FUNCTION_BLOCK "FB_CrossCutsModbus_V1.00"   // FB1, LAD
TITLE = Cross cut machine V1.00
{ S7_Optimized_Access := 'TRUE' }
VERSION : 0.1
   VAR_INPUT
      IN_dMachineIndex : DInt;   // Tracking machine index
      IN_dGlassBreakMachineIndex : DInt;   // Glass break machine index
      IN_dGlassSearchMachineIndex_Q0 : DInt;   // Glass search machine index
      IN_dGlassSearchMachineIndex_Q1 : DInt;   // Glass search machine index
      IN_dGlassSearchMachineIndex_Q2 : DInt;   // Glass search machine index
      IN_dGlassSearchMachineIndex_Q3 : DInt;   // Glass search machine index
      IN_dXCutIndex : DInt;   // Index of the XCUT (0=XC#1, 1=XC#2...)
      IN_xCycleON : Bool;   // Cycle ON
      IN_xGeneralReset : Bool;   // General reset
      IN_xResetAlarms : Bool;   // Reset alarms
      IN_xFaultsEnabled : Bool;   // Faults enabled
      IN_xSimulationActive : Bool;   // Enable simulation (EXPERT USER)
      IN_xMBDone : Bool;   // Modbus client done
      IN_xMBError : Bool;   // Xcut DB
   END_VAR
   VAR_IN_OUT
      INO_tTrack : "UDT_CapData_Tracking";   // Tracking plate
      INO_tEnc : "UDT_Encoder";   // Encoder data
      INO_tOBInit : "GP_OB_Initialize";   // OB Initialize
      INO_tRibbon : "UDT_RibbonData";   // Ribbon data
      INO_tXCutOpt : "FB_CrossCutOpt_V1.00";   // Ribbon data
   END_VAR
   VAR RETAIN
      tHMW : Struct   // HMI Write data
         xCutBreakEnabled : Bool;   // Cut on glass break enabled {X|X|X|X|O}
         xUpdateDistSnap : Bool;   // Update distance from snap roll {X|X|X|X|M}
         xUpdateAngleValue : Bool;   // Update angle value {X|X|X|X|M}
         xIncAngleValue : Bool;   // Increment angle value {X|X|X|X|O}
         xDecAngleValue : Bool;   // Decrement angle value {X|X|X|X|O}
         xUpdateDistCenterLine : Bool;   // Update distance from center line {X|X|X|X|M}
         xCalibDistRequest : Bool;   // Calibration distance request {X|X|X|X|O}
         xCalibDiagRequest : Bool;   // Calibration diagonal request {X|X|X|X|O}
         tManCmd : Struct   // Manual command
            xMan_JogForward : Bool;   // Manual mode - Jog forward {X|X|X|X|M}
            xMan_JobBackward : Bool;   // Manual mode - Jog backward {X|X|X|X|M}
            xMan_CarriageDown : Bool;   // Manual mode - Carriage down {X|X|X|X|M}
            xMan_FireOn : Bool;   // Manual mode - Fire ON {X|X|X|X|M}
            xMan_OilOn : Bool;   // Manual mode - Oil ON {X|X|X|X|M}
         END_STRUCT;
         xCutOperator : Bool;   // Cutting position by operator request {X|X|X|X|O}
         xCutGross : Bool;   // Cutting position by gross width position {X|X|X|X|O}
         xCutNet : Bool;   // Cutting position by net width position {X|X|X|X|O}
         xCutYCut : Bool;   // Cutting position by YCut position {X|X|X|X|O}
         dOperStartCutPos_cmm : DInt;   // Operator start cut position [mm/100] {mm/100|mm|-3000|0|O}
         dOperEndCutPos_cmm : DInt;   // Operator end cut position [mm/100] {mm/100|mm|0|3000|O}
         dDescReactTime_ms : DInt;   // Carriage descent reaction time [ms] {ms|s|0|1|M}
         dRaiseReactTime_ms : DInt;   // Carriage raise reaction time [ms] {ms|s|0|1|M}
         dFireONReactTime_ms : DInt;   // Fire ON reaction time [ms] {ms|s|0|1|M}
         dFireOFFReactTime_ms : DInt;   // Fire OFF reaction time [ms] {ms|s|0|1|M}
         dOilONDelay_ms : DInt;   // Oil ON delay [ms] {ms|s|-1|1|O}
         dOilOFFDelay_ms : DInt;   // Oil OFF delay [ms] {ms|s|-1|1|O}
         dCutStartOffsetDelay_cmm : DInt;   // Start cut offset delay [mm/100] {mm/100|mm|-500|500|O}
         dCutEndOffsetDelay_cmm : DInt;   // End cut offset delay [mm/100] {mm/100|mm|-500|500|O}
         dDistanceFromSnaproll_cmm : DInt;   // Distance from snaproll [mm/100] {mm/100|mm|0|10000|M}
         dAngleValue_uDegree : DInt;   // Bridge angle value [°/1000000] {°/1000000|°|7|9|M}
         dDistanceFromCenterLine_cmm : DInt;   // Distance from center line [mm/100] {mm/100|mm|-3000|0|M}
         dDistTeoLength_cmm : DInt;   // Calibration distance.Theorical length [mm/100] {mm/100|mm|0|7000|O}
         dDistRealLength_cmm : DInt;   // Calibration distance.Real length [mm/100] {mm/100|mm|0|7000|O}
         dDiagRealLength_cmm : DInt;   // Calibration diagonal.Real length [mm/100] {mm/100|mm|0|7000|O}
         dDiagRealWidth_cmm : DInt;   // Calibration diagonal.Real width [mm/100] {mm/100|mm|0|4000|O}
         dDiagGlassFlow_cmm : DInt;   // Calibration diagonal.Real length diagonal glass flow [mm/100] {mm/100|mm|0|10000|O}
         dDiagGlassOppFlow_cmm : DInt;   // Calibration diagonal.Real length diagonal opposite glass flow [mm/100] {mm/100|mm|0|10000|O}
         dCuttingPressure_mN : DInt;   // Cutting pressure [N/1000] {N/1000|N|9|180|O}
         dPosOffset_cmm : DInt;   // Calibration offset distance from snaproll [mm/100] {mm/100|mm|-50|50|O}
         dCutPriority : DInt;   // Cut priority number {X|X|0|5|O}
         xResetHeadUsage : Bool;   // Reset the head usage {X|X|X|X|O}
         xEnDisManCom : Bool;   // Enable disable manual command {X|X|X|X|M}
      END_STRUCT;
      tHMR : Struct   // HMI Read data
         tManCmd : Struct   // Manual command
            xManJogFwdFdbk : Bool;   // Manual jog forward feedback {X|X|X|X|O}
            xManJogBckFdbk : Bool;   // Manual jog backward feedback {X|X|X|X|O}
            xManCarriageDownFdbk : Bool;   // Manual carriage down feedback {X|X|X|X|O}
            xManFireONFdbk : Bool;   // Manual fire ON feedback {X|X|X|X|O}
            xManOilONFdbk : Bool;   // Manual oil ON feedback {X|X|X|X|O}
         END_STRUCT;
         dActualCutPosRequest : DInt;   // Actual cut position request (1=By operator 2=On gross ribbon 3=On net ribbon 4=On YCut position) {X|X|X|X|O}
         dXCutStatusRequest : DInt;   // XCut status request (1=Disabled 3=Enabled) {X|X|X|X|O}
         dXCutActualStatus : DInt;   // XCut actual status (1=Disabled 3=Enabled) {X|X|X|X|O}
         dDistanceFromSnaproll_cmm : DInt;   // Distance from snaproll [mm/100] {mm/100|mm|X|X|O}
         dAngleValue_uDegree : DInt;   // Angle value [°/1000000] {°/1000000|°|X|X|O}
         dDistanceFromCenterLine_cmm : DInt;   // Distance from center line [mm/100] {mm/100|mm|X|X|O}
         dCarriagePosition_cmm : DInt;   // Actual carriage position [mm/100]
         dStatus : DInt;   // XCut actual status (1=Idle 3=Running 7=Faulted) {X|X|X|X|O}
         rHeadUsage_km : Real;   // Head usage [Km] {Km|Km|X|X|O}
         xManComEn : Bool;   // Manual command enabled {X|X|X|X|O}
         dTimeHeadDown_ms : DInt;   // Time head down [ms] {ms|s|X|X|O}
      END_STRUCT;
   END_VAR
   VAR
      tALM : Struct   // HMI Alarms
         tE : Struct   // Emergency alarms
            xLocON : Bool;   // KE.Local emergency ON {X|X|X|X|O}
            xLocal1 : Bool;   // SB.Local emergency push button 1 {X|X|X|X|O}
            xLocal2 : Bool;   // SB.Local emergency push button 2 {X|X|X|X|O}
            xLocal3 : Bool;   // SB.Local emergency push button 3 {X|X|X|X|O}
            xSpare_4 : Bool;
            xSpare_5 : Bool;
            xSpare_6 : Bool;
            xSpare_7 : Bool;
            xSpare_8 : Bool;
            xSpare_9 : Bool;
            xSpare_10 : Bool;
            xSpare_11 : Bool;
            xSpare_12 : Bool;
            xSpare_13 : Bool;
            xSpare_14 : Bool;
            xSpare_15 : Bool;
            xSpare_16 : Bool;
            xSpare_17 : Bool;
            xSpare_18 : Bool;
            xSpare_19 : Bool;
            xSpare_20 : Bool;
            xSpare_21 : Bool;
            xSpare_22 : Bool;
            xSpare_23 : Bool;
            xSpare_24 : Bool;
            xSpare_25 : Bool;
            xSpare_26 : Bool;
            xSpare_27 : Bool;
            xSpare_28 : Bool;
            xSpare_29 : Bool;
            xSpare_30 : Bool;
            xSpare_31 : Bool;
         END_STRUCT;
         tS : Struct   // Stopping faults
            xAxisNotAvail : Bool;   // AZ.Axis not available {X|X|X|X|O}
            xInpInstallation : Bool;   // L+.Input power supply ON {X|X|X|X|O}
            xAuxPower : Bool;   // L+.Auxiliary power supple set-in {X|X|X|X|O}
            xAreaSafety : Bool;   // KE.Area safety {X|X|X|X|O}
            xOverstroke : Bool;   // KA.Carriage overstroke {X|X|X|X|O}
            xExternInputPower : Bool;   // L+.External input power supply {X|X|X|X|O}
            xCarriageCutOut : Bool;   // QM.Carriage translation overload {X|X|X|X|O}
            xDriveTrip : Bool;   // AZ.Drive trip {X|X|X|X|O}
            xDriveNotEnabled : Bool;   // AZ.Drive not enabled {X|X|X|X|O}
            xAxisNotReady : Bool;   // AZ.Axis not ready {X|X|X|X|O}
            xDriveNotReady : Bool;   // AZ.Drive not ready {X|X|X|X|O}
            xAxisNotSyncro : Bool;   // AZ.Axis not syncronized {X|X|X|X|O}
            xSpare_12 : Bool;
            xSpare_13 : Bool;
            xSpare_14 : Bool;
            xSpare_15 : Bool;
            xSpare_16 : Bool;
            xSpare_17 : Bool;
            xSpare_18 : Bool;
            xSpare_19 : Bool;
            xSpare_20 : Bool;
            xSpare_21 : Bool;
            xSpare_22 : Bool;
            xSpare_23 : Bool;
            xSpare_24 : Bool;
            xSpare_25 : Bool;
            xSpare_26 : Bool;
            xSpare_27 : Bool;
            xSpare_28 : Bool;
            xSpare_29 : Bool;
            xSpare_30 : Bool;
            xSpare_31 : Bool;
         END_STRUCT;
         tF : Struct   // Faults
            xSpare_0 : Bool;
            xSpare_1 : Bool;
            xSpare_2 : Bool;
            xSpare_3 : Bool;
            xSpare_4 : Bool;
            xSpare_5 : Bool;
            xSpare_6 : Bool;
            xSpare_7 : Bool;
            xSpare_8 : Bool;
            xSpare_9 : Bool;
            xSpare_10 : Bool;
            xSpare_11 : Bool;
            xSpare_12 : Bool;
            xSpare_13 : Bool;
            xSpare_14 : Bool;
            xSpare_15 : Bool;
            xSpare_16 : Bool;
            xSpare_17 : Bool;
            xSpare_18 : Bool;
            xSpare_19 : Bool;
            xSpare_20 : Bool;
            xSpare_21 : Bool;
            xSpare_22 : Bool;
            xSpare_23 : Bool;
            xSpare_24 : Bool;
            xSpare_25 : Bool;
            xSpare_26 : Bool;
            xSpare_27 : Bool;
            xSpare_28 : Bool;
            xSpare_29 : Bool;
            xSpare_30 : Bool;
            xSpare_31 : Bool;
         END_STRUCT;
         tW : Struct   // Warnings
            xSpare_0 : Bool;
            xSpare_1 : Bool;
            xSpare_2 : Bool;
            xSpare_3 : Bool;
            xSpare_4 : Bool;
            xSpare_5 : Bool;
            xSpare_6 : Bool;
            xSpare_7 : Bool;
            xSpare_8 : Bool;
            xSpare_9 : Bool;
            xSpare_10 : Bool;
            xSpare_11 : Bool;
            xSpare_12 : Bool;
            xSpare_13 : Bool;
            xSpare_14 : Bool;
            xSpare_15 : Bool;
            xSpare_16 : Bool;
            xSpare_17 : Bool;
            xSpare_18 : Bool;
            xSpare_19 : Bool;
            xSpare_20 : Bool;
            xSpare_21 : Bool;
            xSpare_22 : Bool;
            xSpare_23 : Bool;
            xSpare_24 : Bool;
            xSpare_25 : Bool;
            xSpare_26 : Bool;
            xSpare_27 : Bool;
            xSpare_28 : Bool;
            xSpare_29 : Bool;
            xSpare_30 : Bool;
            xSpare_31 : Bool;
         END_STRUCT;
      END_STRUCT;
      ST_xPhaseInProgress : Bool;   // Phases are in progress
      AUX_xValidUpCap : Bool;   // Upstream cap is valid
      AUX_xValidDwCap : Bool;   // Downstream cap is valid
      AUX_dUpCapIndex : DInt;   // Index of the upstream cap
      AUX_dDwCapIndex : DInt;   // Index of the downstream cap
      OS_xNewCapUp : Bool;   // New cap arrived upstream
      OS_xNewCapDw : Bool;   // New cap arrived downstream
      OS_xNewCap : Bool;   // New cap arrived
      ST_xStoppingFaults : Bool;   // Stopping faults
      ST_xFaults : Bool;   // Faults
      ST_xWarnings : Bool;   // Warnings
      ST_xOutputEnabled : Bool;   // Output enabled
      ST_xGlassBreak : Bool;   // Glass break under bridge
      ST_xQualitWithFixedXcut : Bool;   // Quality cap with fixed xcut choice coming
      AUX_dCutStartPosUp_cmm : DInt;   // Cut start position upstream [mm/100]
      AUX_dCutStopPosUp_cmm : DInt;   // Cut stop position downstream [mm/100]
      AUX_dCutStartPosDw_cmm : DInt;   // Cut start position downstream [mm/100]
      AUX_dCutStopPosDw_cmm : DInt;   // Cut stop position downstream [mm/100]
      AUX_xUpIsQuality : Bool;   // Upstream cap is a quality cap
      AUX_xDwIsQuality : Bool;   // Downstream cap is a quality cap
      PH_xCutRequest : Bool;   // Cut request phase
      PH_xWriteModbus : Bool;   // Modbus write phase
      PH_xEndWriteModbus : Bool;   // Modbus end write phase
      PH_xReadModbus : Bool;   // Modbus read phase
      PH_xEndReadModbus : Bool;   // Modbus end read phase
      AUX_dMissionCounterValue_cmm : DInt;   // Mission counter value to inverter [mm/100]
      AUX_dMissionToSend : DInt;   // Index mission send to inverter
      AUX_tOutputDrive : "UDT_XCUT_DRIVE_OUTPUT";   // Copy of output area drive
      PH_xEndCutRequest : Bool;   // End cut request phase
      OSR_xButtonEnabled : Bool;   // OSR.Button enabled
      OS_xButtonEnabled : Bool;   // OS.Button enabled
      AUX_dLastLiveCounter : DInt;
      tmON_InvCoutTimeout : TON_TIME;   // Inverter counter timeout
      tmON_AxisSyncroTimeout : TON_TIME;   // Inverter counter timeout
      AUX_dNextPlateTime_ms : DInt;   // Next plate arriving time [ms]
      AUX_dCutTime20Per_ms : DInt;   // Cutting time at 20 percent [ms]
      AUX_dCutTime40Per_ms : DInt;   // Cutting time at 40 percent [ms]
      AUX_dCutTime60Per_ms : DInt;   // Cutting time at 60 percent [ms]
      AUX_dCutTime80Per_ms : DInt;   // Cutting time at 80 percent [ms]
      AUX_dCutTime100Per_ms : DInt;   // Cutting time at 100 percent [ms]
      ST_xCondOkMan : Bool;   // Condition ok manual command
      AUX_dSimWaitEnd_ms : DInt;   // Simulation waiting end cut [ms]
      AUX_dSimCutTime_ms : DInt;   // Simulation cutting time [ms]
      AUX_dSimCutSpace_cmm : DInt;   // Simulation cutting space [mm/100]
      AUX_dSimStoreCutTime_ms : DInt;   // Simulation saved cutting time [ms]
      AUX_rgdParameterArray : Array[0..39] of DInt;   // Array of xcut parameters (menu 20)
      AUX_rgtIN_tDriveData : "UDT_XCUT_DRIVE_INPUT";   // Drive input data
      AUX_rgtOUT_tDriveData : "UDT_XCUT_DRIVE_OUTPUT";   // Drive output data
   END_VAR
   VAR_TEMP
      TMP_rValue : LReal;   // Temp real value
      TMP_xCalcMission : Bool;   // Temp calculate mission
      TMP_dwValue : DWord;   // Temp Dint value
      TMP_dValue : DInt;   // Temp Dint value
      TMP_xUpdateKM : Bool;   // OS update KM counter
      TMP_dCutTime_ms : DInt;   // Cut time [ms]
      TMP_dConstTime_ms : DInt;   // Const time [ms]
      TMP_rAccTime_s : Real;   // Acceleration time [ms]
      TMP_dTravSpace_cmm : DInt;   // Travel space [mm/100]
      TMP_dCutSpace_cmm : DInt;   // Cut Space [mm/100]
      TMP_dCutYSpace_cmm : DInt;   // Cut y space [mm/100]
      TMP_dConstSpace_cmm : DInt;   // Const space [mm/100]
      TMP_dRampSpace_cmm : DInt;   // Ramp space [mm/100]
      TMP_dRetVal : DInt;   // Ramp space [mm/100]
      TMP_rDiagGlassFlow_cmm : Real;
      TMP_rDiagRealWidth_cmm : Real;
      TMP_rDiagRealLength_cmm : Real;
      TMP_iModbus_mode : UDInt;   // Modbus mode (0=read, 1=write)
      TMP_dModbus_address : UDInt;   // Modbus address
      TMP_dModbus_length : UDInt;   // Modbus data length
      TMP_vDataPointer : Variant;
      TMP_dIndex : DInt;
   END_VAR
   VAR CONSTANT
      CONST_DREACTTIMETRACK_MS : DInt := 50;   // Tracking machine reaction time [ms]
      CONST_DMODECUT_OPERATOR : DInt := 1;   // Cut modality - By operator
      CONST_DMODECUT_GROSS : DInt := 2;   // Cut modality - Gross width
      CONST_DMODECUT_NET : DInt := 3;   // Cut modality - Net width
      CONST_DMODECUT_YCUT : DInt := 4;   // Cut modality - YCut
      CONST_DMINCUTRANGE_CMM : DInt := 25000;   // Minimum cutting start position [mm/100]
      CONST_DMAXCUTRANGE_CMM : DInt := 500000;   // Maximum cutting start position [mm/100]
      CONST_DMAXMISSIONNUM : DInt := 1000;   // Maximum number of mission to XCUT
      CONST_DMAXWAITFEEDBACK_CMM : DInt := 20000;   // Waiting space feedback [mm/100]
      CONST_DDISABLED : DInt := 1;   // Disabled
      CONST_DENABLED : DInt := 3;   // Enabled
      CONST_DSIZEALARMS : UDInt := 32;   // Number of bool on alarms structure
      CONST_DTIMEOUTINVERTER_MS : Time := T#2000ms;   // Inverter counter timeout
      CONST_DMAXRETSPEED_RPM : DInt := 3750;   // Maximum return speed [rpm]
      CONST_DSPEED_CMM_S : DInt := 500000;   // Return travel speed [mm/100/s]
      CONST_DRAMP_CMM_S2 : DInt := 1200000;   // Return travel ramp [mm/100/s]
      CONST_DBREAKDOWNOFF_CMM : DInt := 50000;   // Break downstream offset [mm/100]
      CONST_DBREAKUPOFF_CMM : DInt := 50000;   // Break upstream offset [mm/100]
      CONST_DADDRESSMENU_READ : UDInt := 2001;   // Parameter menu start (#20.01=2001)
      CONST_DADDRESSMENU_WRITE : UDInt := 2010;   // Parameter menu start (#20.01=2001)
      CONST_DSEARCHQLTUPSTREAM_CMM : DInt := 1000000;   // Search qlt cap upstream limit [mm/100]
      CONST_DSEARCHQLTDOWNSTREAM_CMM : DInt := 400000;   // Search qlt cap downstream limit [mm/100]
   END_VAR
   VAR_TEMP   // added for the SCL form of the ladder/FBD networks
      _w1 : Bool;
   END_VAR
   // // AUX_rgdParameterArray[0] : #20.01
   // // AUX_rgdParameterArray[1] : #20.02
   // // AUX_rgdParameterArray[2] : #20.03
   // // AUX_rgdParameterArray[3] : #20.04
   // // AUX_rgdParameterArray[4] : #20.05
   // // AUX_rgdParameterArray[5] : #20.06
   // // AUX_rgdParameterArray[6] : #20.07
   // // AUX_rgdParameterArray[7] : #20.08
   // // AUX_rgdParameterArray[8] : #20.09
   // // AUX_rgdParameterArray[9] : #20.10
   // // AUX_rgdParameterArray[10] : #20.11
   // // AUX_rgdParameterArray[11] : #20.12
   // // AUX_rgdParameterArray[12] : #20.13
   // // AUX_rgdParameterArray[13] : #20.14
   // // AUX_rgdParameterArray[14] : #20.15
   // // AUX_rgdParameterArray[15] : #20.16
   // // AUX_rgdParameterArray[16] : #20.17
   // // AUX_rgdParameterArray[17] : #20.18
   // // AUX_rgdParameterArray[18] : #20.19
   // // AUX_rgdParameterArray[19] : #20.20
   // // AUX_rgdParameterArray[20] : #20.21
   // // AUX_rgdParameterArray[21] : #20.22
   // // AUX_rgdParameterArray[22] : #20.23
   // // AUX_rgdParameterArray[23] : #20.24
   // // AUX_rgdParameterArray[24] : #20.25
   // // AUX_rgdParameterArray[25] : #20.26
   // // AUX_rgdParameterArray[26] : #20.27
   // // AUX_rgdParameterArray[27] : #20.28
   // // AUX_rgdParameterArray[28] : #20.29
   // // AUX_rgdParameterArray[29] : #20.30
   // // AUX_rgdParameterArray[30] : #20.31
   // // AUX_rgdParameterArray[31] : #20.32
   // // AUX_rgdParameterArray[32] : #20.33
   // // AUX_rgdParameterArray[33] : #20.34
   // // AUX_rgdParameterArray[34] : #20.35
   // // AUX_rgdParameterArray[35] : #20.36
   // // AUX_rgdParameterArray[36] : #20.37
   // // AUX_rgdParameterArray[37] : #20.38
   // // AUX_rgdParameterArray[38] : #20.39
   // // AUX_rgdParameterArray[39] : #20.40
BEGIN

REGION Network 1: ####_CONSTANTS_####
END_REGION

REGION Network 2: ####_MATCH_####
END_REGION

REGION Network 3 (SCL): Update data from inverter
   IF #PH_xEndReadModbus THEN

   #AUX_rgtIN_tDriveData.dCarriagePos_dmm := #AUX_rgdParameterArray[30];
   #AUX_rgtIN_tDriveData.dLehrPosition_cmm := #AUX_rgdParameterArray[32];
   #AUX_rgtIN_tDriveData.dLehrSpeed_cmm_min := #AUX_rgdParameterArray[36];
   #AUX_rgtIN_tDriveData.dErrorCode := #AUX_rgdParameterArray[34];
   #AUX_rgtIN_tDriveData.dMissionDone := #AUX_rgdParameterArray[35];
   #AUX_rgtIN_tDriveData.dMissionUnDone := #AUX_rgdParameterArray[33];
   #AUX_rgtIN_tDriveData.iLiveCounter := DINT_TO_INT(#AUX_rgdParameterArray[9]);
   #AUX_rgtIN_tDriveData.iTimeHeadDown_ms := DINT_TO_INT(#AUX_rgdParameterArray[10]);
   #TMP_dwValue := DINT_TO_DWORD(#AUX_rgdParameterArray[29]);
   SCATTER(IN:=#TMP_dwValue,
           OUT=>#AUX_rgtIN_tDriveData.rgxStatusBits);

   #PH_xEndReadModbus := 0;
   END_IF;
END_REGION

REGION Network 4 (SCL): General reset
   IF #IN_xGeneralReset THEN

       #PH_xCutRequest := FALSE;
       #PH_xEndCutRequest := FALSE;
       #AUX_xValidDwCap := FALSE;
       #AUX_xValidUpCap := FALSE;

   END_IF;
END_REGION

REGION Network 5 (SCL): Move data information to tracking
   #INO_tTrack.rgtTrackMachine[#IN_dMachineIndex].tUserData.dSetDistanceSnap_cmm := #tHMR.dDistanceFromSnaproll_cmm + #tHMW.dPosOffset_cmm + 10000; //100mm is an offset fixed value
   #INO_tTrack.rgtTrackMachine[#IN_dMachineIndex].tUserData.dSetMachReacTime_ms := #CONST_DREACTTIMETRACK_MS;
END_REGION

REGION Network 6 (SCL): Manage tracking call

   #OS_xNewCapUp := FALSE;
   #OS_xNewCapDw := FALSE;
   #OS_xNewCap := FALSE;

   IF #INO_tTrack.rgtTrackMachine[#IN_dMachineIndex].tUserData.xGetPosReach THEN

       #AUX_xUpIsQuality := FALSE;
       #AUX_xDwIsQuality := FALSE;

       IF (NOT #ST_xPhaseInProgress) THEN

           #OS_xNewCap := TRUE;

           IF #INO_tTrack.rgtTrackMachine[#IN_dMachineIndex].tUserData.dGetUpstremIndex >= 0 THEN
               #AUX_xValidUpCap := TRUE;
               #OS_xNewCapUp := TRUE;            
               #AUX_dUpCapIndex := #INO_tTrack.rgtTrackMachine[#IN_dMachineIndex].tUserData.dGetUpstremIndex;

               //Evaluate if is a quality plate
               IF  #INO_tTrack.rgtTrackCaps[#AUX_dUpCapIndex].tCap.rgtLites[0].dMainDestination = "DQUALITYDESTMASK1" OR
                   #INO_tTrack.rgtTrackCaps[#AUX_dUpCapIndex].tCap.rgtLites[0].dMainDestination = "DQUALITYDESTMASK2" OR
                   #INO_tTrack.rgtTrackCaps[#AUX_dUpCapIndex].tCap.rgtLites[0].dMainDestination = "DQUALITYDESTMASK3" OR
                   #INO_tTrack.rgtTrackCaps[#AUX_dUpCapIndex].tCap.rgtLites[0].dMainDestination = "DQUALITYDESTMASK4" THEN

                  #AUX_xUpIsQuality := TRUE;

               END_IF;

           ELSE
               #AUX_xValidUpCap := FALSE;
               #OS_xNewCapUp := FALSE;            
               #AUX_dUpCapIndex := 0;
           END_IF;

           IF #INO_tTrack.rgtTrackMachine[#IN_dMachineIndex].tUserData.dGetDownstreamIndex >= 0 THEN
               #AUX_xValidDwCap := TRUE;
               #OS_xNewCapDw := TRUE;            
               #AUX_dDwCapIndex := #INO_tTrack.rgtTrackMachine[#IN_dMachineIndex].tUserData.dGetDownstreamIndex;

               //Evaluate if is a quality plate
               IF  #INO_tTrack.rgtTrackCaps[#AUX_dDwCapIndex].tCap.rgtLites[0].dMainDestination = "DQUALITYDESTMASK1" OR
                   #INO_tTrack.rgtTrackCaps[#AUX_dDwCapIndex].tCap.rgtLites[0].dMainDestination = "DQUALITYDESTMASK2" OR
                   #INO_tTrack.rgtTrackCaps[#AUX_dDwCapIndex].tCap.rgtLites[0].dMainDestination = "DQUALITYDESTMASK3" OR
                   #INO_tTrack.rgtTrackCaps[#AUX_dUpCapIndex].tCap.rgtLites[0].dMainDestination = "DQUALITYDESTMASK4" THEN

                  #AUX_xDwIsQuality := TRUE;

               END_IF;

           ELSE
               #AUX_xValidDwCap := FALSE;
               #OS_xNewCapDw := FALSE;            
               #AUX_dDwCapIndex := 0;
           END_IF;



       END_IF;

       #INO_tTrack.rgtTrackMachine[#IN_dMachineIndex].tUserData.xGetPosReach := FALSE;

   END_IF;
END_REGION

REGION Network 7: OS enable disable XCut buttons
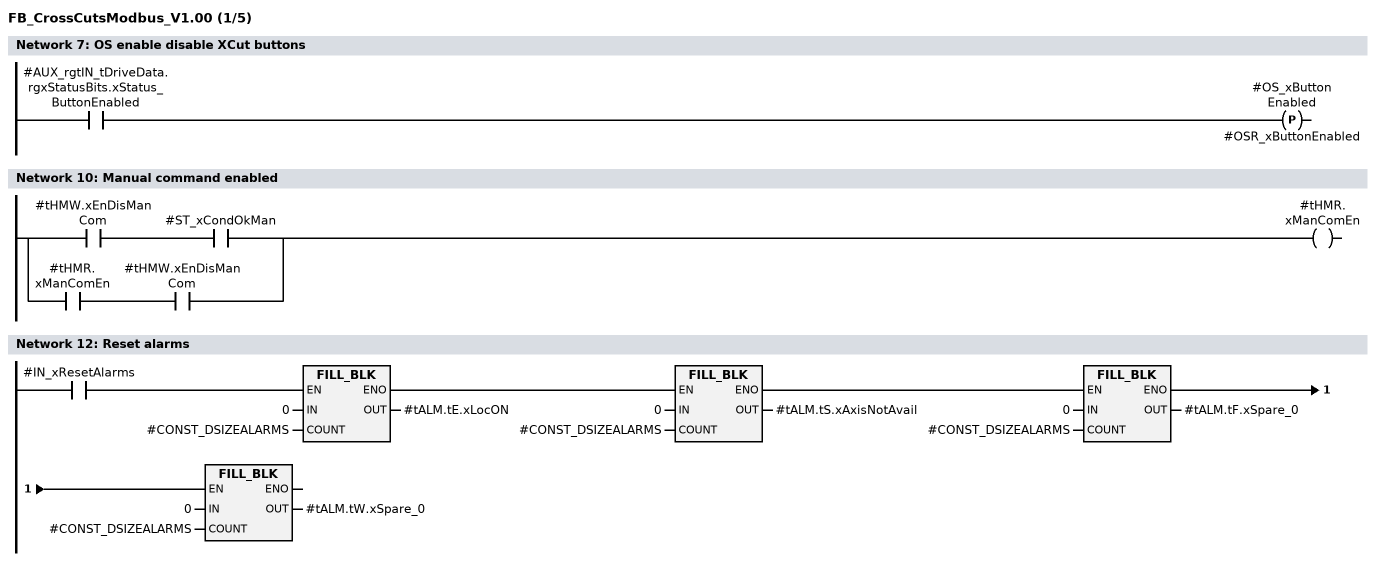
   #OS_xButtonEnabled := #AUX_rgtIN_tDriveData.rgxStatusBits.xStatus_ButtonEnabled AND NOT #OSR_xButtonEnabled;   // rising edge
   #OSR_xButtonEnabled := #AUX_rgtIN_tDriveData.rgxStatusBits.xStatus_ButtonEnabled;
END_REGION

REGION Network 8: ####_HMI_LOGICS_####
END_REGION

REGION Network 9 (SCL): List of HMI logics
   REGION UpdateDistanceSnaproll

   IF #tHMW.xUpdateDistSnap THEN
       #tHMW.xUpdateDistSnap := FALSE;

       #tHMR.dDistanceFromSnaproll_cmm := #tHMW.dDistanceFromSnaproll_cmm;

   END_IF;

   END_REGION

   REGION UpdateAngleValue

   IF #tHMW.xUpdateAngleValue THEN
       #tHMW.xUpdateAngleValue := FALSE;

       #tHMR.dAngleValue_uDegree := #tHMW.dAngleValue_uDegree;

   END_IF;

   END_REGION

   REGION UpdateDistanceCenterLine

   IF #tHMW.xUpdateDistCenterLine THEN
       #tHMW.xUpdateDistCenterLine := FALSE;

       #tHMR.dDistanceFromCenterLine_cmm := #tHMW.dDistanceFromCenterLine_cmm;

   END_IF;

   END_REGION
   (* REGION EnableDisableCutOnBreak

   IF #tHMW.xEnCutBreak THEN    
       #tHMW.xEnCutBreak := FALSE;
       #tHMR.xCutBreakEnabled := TRUE;
   END_IF;

   IF #tHMW.xDisCutBreak THEN    
       #tHMW.xDisCutBreak := FALSE;
       #tHMR.xCutBreakEnabled := FALSE;
   END_IF;

   END_REGION *)

   (* REGION EnableDisableCut

   IF #tHMW.xEnableCut OR (#tHMR.dXCutStatusRequest = #CONST_DDISABLED AND #OS_xButtonEnabled) THEN    
       #tHMW.xEnableCut := FALSE;
       #tHMR.dXCutStatusRequest := #CONST_DENABLED;
   ELSIF #tHMW.xDisableCut OR (#tHMR.dXCutStatusRequest = #CONST_DENABLED AND #OS_xButtonEnabled) THEN    
       #tHMW.xDisableCut := FALSE;
       #tHMR.dXCutStatusRequest := #CONST_DDISABLED;
   END_IF;


   END_REGION
   *)
   REGION IncDecAngleValue

       IF #tHMW.xIncAngleValue THEN
           #tHMW.xIncAngleValue := FALSE;
           #tHMR.dAngleValue_uDegree := #tHMR.dAngleValue_uDegree + 10000;
           #tHMW.dAngleValue_uDegree := #tHMR.dAngleValue_uDegree;
       END_IF;

   IF #tHMW.xDecAngleValue THEN
       #tHMW.xDecAngleValue := FALSE;
       #tHMR.dAngleValue_uDegree := #tHMR.dAngleValue_uDegree - 10000;
       #tHMW.dAngleValue_uDegree := #tHMR.dAngleValue_uDegree;

   END_IF;

   END_REGION

   REGION DistanceCalibration

   IF #tHMW.xCalibDistRequest THEN

       #tHMW.xCalibDistRequest := FALSE;

       #tHMR.dDistanceFromSnaproll_cmm := #tHMW.dDistRealLength_cmm - #tHMW.dDistTeoLength_cmm + #tHMR.dDistanceFromSnaproll_cmm;

   END_IF;   

   END_REGION

   REGION DiagonalCalibration

   IF #tHMW.xCalibDiagRequest THEN

       #tHMW.xCalibDiagRequest := FALSE;
       #TMP_rDiagGlassFlow_cmm := DINT_TO_REAL(#tHMW.dDiagGlassFlow_cmm);
       #TMP_rDiagRealWidth_cmm := DINT_TO_REAL(#tHMW.dDiagRealWidth_cmm);
       #TMP_rDiagRealLength_cmm := DINT_TO_REAL(#tHMW.dDiagRealLength_cmm);

       #TMP_rValue := (((ATAN((SQRT(#TMP_rDiagGlassFlow_cmm**2 - #TMP_rDiagRealWidth_cmm**2) - #TMP_rDiagRealLength_cmm) / #TMP_rDiagRealWidth_cmm) * 360.0) / 2.0) / 3.141593) * 1000000.0;
       #tHMR.dAngleValue_uDegree := #tHMR.dAngleValue_uDegree + LREAL_TO_DINT(#TMP_rValue);

   END_IF;   

   END_REGION

   REGION Cutting position request

   IF #tHMW.xCutOperator THEN
       #tHMW.xCutOperator := FALSE;
       #tHMR.dActualCutPosRequest := #CONST_DMODECUT_OPERATOR;
   END_IF;    

   IF #tHMW.xCutGross THEN
       #tHMW.xCutGross := FALSE;
       #tHMR.dActualCutPosRequest := #CONST_DMODECUT_GROSS;
   END_IF;    

   IF #tHMW.xCutNet THEN
       #tHMW.xCutNet := FALSE;
       #tHMR.dActualCutPosRequest := #CONST_DMODECUT_NET;
   END_IF;    

   IF #tHMW.xCutYCut THEN
       #tHMW.xCutYCut := FALSE;
       #tHMR.dActualCutPosRequest := #CONST_DMODECUT_YCUT;
   END_IF;    

   END_REGION

   REGION Reset head usage

   IF #tHMW.xResetHeadUsage THEN

       #tHMW.xResetHeadUsage := FALSE;

       #tHMR.rHeadUsage_km := 0;
   END_IF;


   END_REGION

   REGION SIMULATION

       IF #IN_xSimulationActive THEN
           #tHMR.dActualCutPosRequest := #CONST_DMODECUT_YCUT;
           #tHMR.dXCutStatusRequest := #CONST_DENABLED;
       END_IF;

   END_REGION
END_REGION

REGION Network 10: Manual command enabled
   RUNG wire#powerrail
      Contact( #tHMW.xEnDisManCom )
      Contact( #ST_xCondOkMan )
      wire#w1
      Coil( #tHMR.xManComEn )
   END_RUNG
   RUNG wire#powerrail
      Contact( #tHMR.xManComEn )
      Contact( #tHMW.xEnDisManCom )
   END_RUNG wire#w1
   // the same network as SCL:
   #tHMR.xManComEn := (#tHMW.xEnDisManCom AND #ST_xCondOkMan) OR (#tHMR.xManComEn AND #tHMW.xEnDisManCom);
END_REGION

REGION Network 11: ####_ALARMS_####
END_REGION

REGION Network 12: Reset alarms
   RUNG wire#powerrail
      Contact( #IN_xResetAlarms )
      FillBlockI(in := 0, count := #CONST_DSIZEALARMS, out => #tALM.tE.xLocON)
      FillBlockI(in := 0, count := #CONST_DSIZEALARMS, out => #tALM.tS.xAxisNotAvail)
      FillBlockI(in := 0, count := #CONST_DSIZEALARMS, out => #tALM.tF.xSpare_0)
      FillBlockI(in := 0, count := #CONST_DSIZEALARMS, out => #tALM.tW.xSpare_0)
   END_RUNG
   // the same network as SCL:
   IF #IN_xResetAlarms THEN
       FILL_BLK(IN := 0, COUNT := #CONST_DSIZEALARMS, OUT => #tALM.tE.xLocON);
       FILL_BLK(IN := 0, COUNT := #CONST_DSIZEALARMS, OUT => #tALM.tS.xAxisNotAvail);
       FILL_BLK(IN := 0, COUNT := #CONST_DSIZEALARMS, OUT => #tALM.tF.xSpare_0);
       FILL_BLK(IN := 0, COUNT := #CONST_DSIZEALARMS, OUT => #tALM.tW.xSpare_0);
   END_IF;
END_REGION

REGION Network 13: Anomaly list
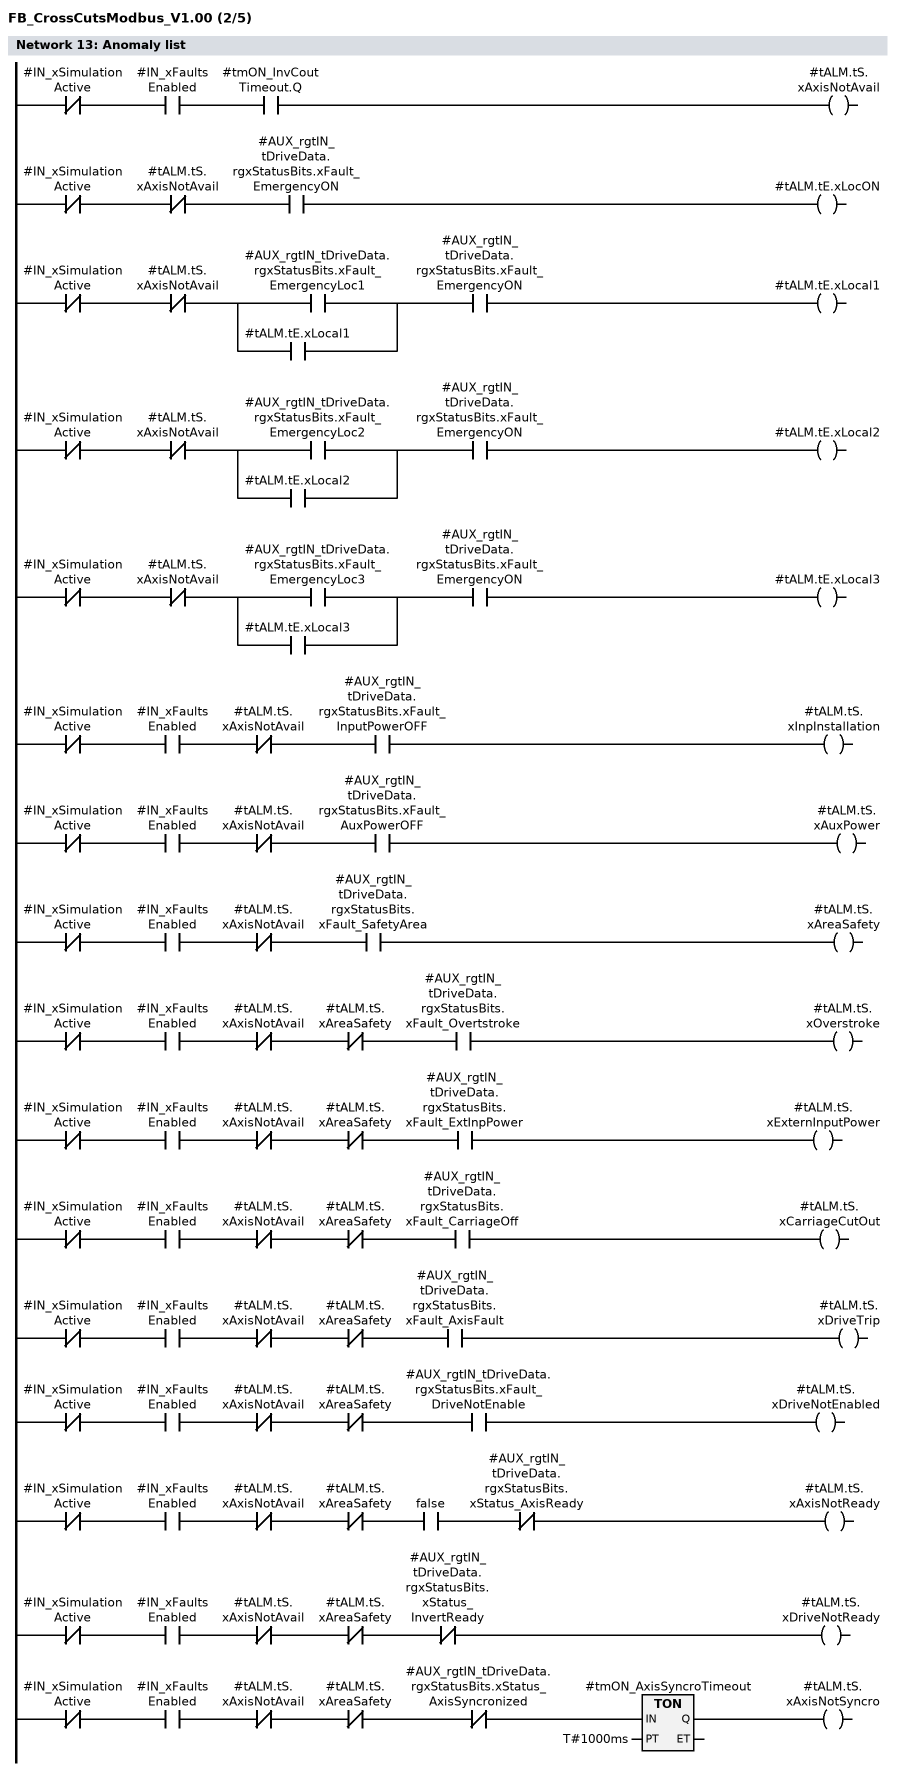
   #tALM.tS.xAxisNotAvail := NOT #IN_xSimulationActive AND #IN_xFaultsEnabled AND #tmON_InvCoutTimeout.Q;
   #tALM.tE.xLocON := NOT #IN_xSimulationActive AND NOT #tALM.tS.xAxisNotAvail AND #AUX_rgtIN_tDriveData.rgxStatusBits.xFault_EmergencyON;
   #tALM.tE.xLocal1 := NOT #IN_xSimulationActive AND NOT #tALM.tS.xAxisNotAvail AND (#AUX_rgtIN_tDriveData.rgxStatusBits.xFault_EmergencyLoc1 OR #tALM.tE.xLocal1) AND #AUX_rgtIN_tDriveData.rgxStatusBits.xFault_EmergencyON;
   #tALM.tE.xLocal2 := NOT #IN_xSimulationActive AND NOT #tALM.tS.xAxisNotAvail AND (#AUX_rgtIN_tDriveData.rgxStatusBits.xFault_EmergencyLoc2 OR #tALM.tE.xLocal2) AND #AUX_rgtIN_tDriveData.rgxStatusBits.xFault_EmergencyON;
   #tALM.tE.xLocal3 := NOT #IN_xSimulationActive AND NOT #tALM.tS.xAxisNotAvail AND (#AUX_rgtIN_tDriveData.rgxStatusBits.xFault_EmergencyLoc3 OR #tALM.tE.xLocal3) AND #AUX_rgtIN_tDriveData.rgxStatusBits.xFault_EmergencyON;
   #tALM.tS.xInpInstallation := NOT #IN_xSimulationActive AND #IN_xFaultsEnabled AND NOT #tALM.tS.xAxisNotAvail AND #AUX_rgtIN_tDriveData.rgxStatusBits.xFault_InputPowerOFF;
   #tALM.tS.xAuxPower := NOT #IN_xSimulationActive AND #IN_xFaultsEnabled AND NOT #tALM.tS.xAxisNotAvail AND #AUX_rgtIN_tDriveData.rgxStatusBits.xFault_AuxPowerOFF;
   #tALM.tS.xAreaSafety := NOT #IN_xSimulationActive AND #IN_xFaultsEnabled AND NOT #tALM.tS.xAxisNotAvail AND #AUX_rgtIN_tDriveData.rgxStatusBits.xFault_SafetyArea;
   #tALM.tS.xOverstroke := NOT #IN_xSimulationActive AND #IN_xFaultsEnabled AND NOT #tALM.tS.xAxisNotAvail AND NOT #tALM.tS.xAreaSafety AND #AUX_rgtIN_tDriveData.rgxStatusBits.xFault_Overtstroke;
   #tALM.tS.xExternInputPower := NOT #IN_xSimulationActive AND #IN_xFaultsEnabled AND NOT #tALM.tS.xAxisNotAvail AND NOT #tALM.tS.xAreaSafety AND #AUX_rgtIN_tDriveData.rgxStatusBits.xFault_ExtInpPower;
   #tALM.tS.xCarriageCutOut := NOT #IN_xSimulationActive AND #IN_xFaultsEnabled AND NOT #tALM.tS.xAxisNotAvail AND NOT #tALM.tS.xAreaSafety AND #AUX_rgtIN_tDriveData.rgxStatusBits.xFault_CarriageOff;
   #tALM.tS.xDriveTrip := NOT #IN_xSimulationActive AND #IN_xFaultsEnabled AND NOT #tALM.tS.xAxisNotAvail AND NOT #tALM.tS.xAreaSafety AND #AUX_rgtIN_tDriveData.rgxStatusBits.xFault_AxisFault;
   #tALM.tS.xDriveNotEnabled := NOT #IN_xSimulationActive AND #IN_xFaultsEnabled AND NOT #tALM.tS.xAxisNotAvail AND NOT #tALM.tS.xAreaSafety AND #AUX_rgtIN_tDriveData.rgxStatusBits.xFault_DriveNotEnable;
   #tALM.tS.xAxisNotReady := NOT #IN_xSimulationActive AND #IN_xFaultsEnabled AND NOT #tALM.tS.xAxisNotAvail AND NOT #tALM.tS.xAreaSafety AND false AND NOT #AUX_rgtIN_tDriveData.rgxStatusBits.xStatus_AxisReady;
   #tALM.tS.xDriveNotReady := NOT #IN_xSimulationActive AND #IN_xFaultsEnabled AND NOT #tALM.tS.xAxisNotAvail AND NOT #tALM.tS.xAreaSafety AND NOT #AUX_rgtIN_tDriveData.rgxStatusBits.xStatus_InvertReady;
   #tmON_AxisSyncroTimeout(IN := NOT #IN_xSimulationActive AND #IN_xFaultsEnabled AND NOT #tALM.tS.xAxisNotAvail AND NOT #tALM.tS.xAreaSafety AND NOT #AUX_rgtIN_tDriveData.rgxStatusBits.xStatus_AxisSyncronized,   // TON
                           PT := T#1000ms);
   #tALM.tS.xAxisNotSyncro := #tmON_AxisSyncroTimeout.Q;
END_REGION

REGION Network 14: ####_STATUSES_####
END_REGION
